screen "BC Max Step Times" 1280x800, template "Template"
   on GenerateScreen: "TitleUpdater"()
   Button "HmiScreenItemData_1" at 1,1 size 150x43; TextOn 'Back'; TextOff 'Commissioning'
      on Release: ActivateScreen("Commissioning Main Page", 0)
   Button "Button_1" at 21,736 size 161x32; TextOff 'Back'
      on Activate: ActivateScreen("IGG Process Times", 0)
   TextField "Text field_25" at 83,285 size 286x22; Text 'Step 040'
   TextField "Text field_29" at 383,118 size 77x20; Text 'Time (ms)'
   TextField "Text field_33" at 83,312 size 286x22; Text 'Step 050'
   IOField "I/O field_58" at 382,312 size 60x22; Authorization "Parameter Change"; FormatPattern s9999999999
      ProcessValue <- "86_Times_STEP_MAX_TIME_STP_050(1)"
   TextField "Text field_35" at 83,367 size 286x22; Text 'Step 070'
   TextField "Text field_65" at 83,144 size 286x22; Text 'Step 001'
   TextField "Text field_67" at 83,173 size 286x22; Text 'Step 005'
   TextField "Text field_69" at 83,200 size 286x22; Text 'Step 010'
   TextField "Text field_71" at 83,229 size 286x22; Text 'Step 020'
   TextField "Text field_73" at 83,257 size 286x22; Text 'Step 030'
   TextField "Text field_42" at 83,118 size 89x20; Text 'Description'
   IOField "I/O field_128" at 382,144 size 60x22; Authorization "Parameter Change"; FormatPattern s9999999999
      ProcessValue <- "86_Times_STEP_MAX_TIME_STP_001(1)"
   IOField "I/O field_133" at 382,173 size 60x22; Authorization "Parameter Change"; FormatPattern s9999999999
      ProcessValue <- "86_Times_STEP_MAX_TIME_STP_005(1)"
   IOField "I/O field_138" at 382,200 size 60x22; Authorization "Parameter Change"; FormatPattern s9999999999
      ProcessValue <- "86_Times_STEP_MAX_TIME_STP_010(1)"
   IOField "I/O field_148" at 382,257 size 60x22; Authorization "Parameter Change"; FormatPattern s9999999999
      ProcessValue <- "86_Times_STEP_MAX_TIME_STP_030(1)"
   IOField "I/O field_64" at 382,367 size 60x22; Authorization "Parameter Change"; FormatPattern s9999999999
      ProcessValue <- "86_Times_STEP_MAX_TIME_STP_070(1)"
   TextField "Text field_53" at 82,92 size 247x26; Text 'BC Maximum Step Times'
   IOField "I/O field_5" at 382,229 size 60x22; Authorization "Parameter Change"; FormatPattern s9999999999
      ProcessValue <- "86_Times_STEP_MAX_TIME_STP_020(1)"
   TextField "Text field_1" at 83,340 size 286x22; Text 'Step 060'
   IOField "I/O field_2" at 382,340 size 60x22; Authorization "Parameter Change"; FormatPattern s9999999999
      ProcessValue <- "86_Times_STEP_MAX_TIME_STP_060(1)"
   TextField "Text field_2" at 461,286 size 286x22; Text 'Step 240'
   TextField "Text field_3" at 750,119 size 77x20; Text 'Time (ms)'
   TextField "Text field_4" at 461,313 size 286x22; Text 'Step 250'
   IOField "I/O field_1" at 758,312 size 60x22; Authorization "Parameter Change"; FormatPattern s9999999999
      ProcessValue <- "86_Times_STEP_MAX_TIME_STP_250(1)"
   TextField "Text field_5" at 461,368 size 286x22; Text 'Step 270'
   TextField "Text field_6" at 461,145 size 286x22; Text 'Step 190'
   TextField "Text field_7" at 461,174 size 286x22; Text 'Step 200'
   TextField "Text field_8" at 461,201 size 286x22; Text 'Step 210'
   TextField "Text field_9" at 461,230 size 286x22; Text 'Step 220'
   TextField "Text field_10" at 461,258 size 286x22; Text 'Step 230'
   TextField "Text field_11" at 461,119 size 89x20; Text 'Description'
   IOField "I/O field_3" at 758,145 size 60x22; Authorization "Parameter Change"; FormatPattern s9999999999
      ProcessValue <- "86_Times_STEP_MAX_TIME_STP_190(1)"
   IOField "I/O field_4" at 758,174 size 60x22; Authorization "Parameter Change"; FormatPattern s9999999999
      ProcessValue <- "86_Times_STEP_MAX_TIME_STP_200(1)"
   IOField "I/O field_6" at 758,201 size 60x22; Authorization "Parameter Change"; FormatPattern s9999999999
      ProcessValue <- "86_Times_STEP_MAX_TIME_STP_210(1)"
   IOField "I/O field_8" at 758,258 size 60x22; Authorization "Parameter Change"; FormatPattern s9999999999
      ProcessValue <- "86_Times_STEP_MAX_TIME_STP_230(1)"
   IOField "I/O field_9" at 758,367 size 60x22; Authorization "Parameter Change"; FormatPattern s9999999999
      ProcessValue <- "86_Times_STEP_MAX_TIME_STP_270(1)"
   IOField "I/O field_10" at 758,230 size 60x22; Authorization "Parameter Change"; FormatPattern s9999999999
      ProcessValue <- "86_Times_STEP_MAX_TIME_STP_220(1)"
   TextField "Text field_13" at 461,341 size 286x22; Text 'Step 260'
   IOField "I/O field_11" at 758,340 size 60x22; Authorization "Parameter Change"; FormatPattern s9999999999
      ProcessValue <- "86_Times_STEP_MAX_TIME_STP_260(1)"
   TextField "Text field_14" at 83,398 size 286x22; Text 'Step 080'
   IOField "I/O field_12" at 382,398 size 60x22; Authorization "Parameter Change"; FormatPattern s9999999999
      ProcessValue <- "86_Times_STEP_MAX_TIME_STP_080(1)"
   TextField "Text field_15" at 83,426 size 286x22; Text 'Step 090'
   IOField "I/O field_13" at 382,426 size 60x22; Authorization "Parameter Change"; FormatPattern s9999999999
      ProcessValue <- "86_Times_STEP_MAX_TIME_STP_090(1)"
   TextField "Text field_16" at 83,453 size 286x22; Text 'Step 100'
   IOField "I/O field_14" at 382,453 size 60x22; Authorization "Parameter Change"; FormatPattern s9999999999
      ProcessValue <- "86_Times_STEP_MAX_TIME_STP_100(1)"
   IOField "I/O field_15" at 382,285 size 60x22; Authorization "Parameter Change"; FormatPattern s9999999999
      ProcessValue <- "86_Times_STEP_MAX_TIME_STP_040(1)"
   TextField "Text field_17" at 461,395 size 286x22; Text 'Step 280'
   IOField "I/O field_16" at 758,394 size 60x22; Authorization "Parameter Change"; FormatPattern s9999999999
      ProcessValue <- "86_Times_STEP_MAX_TIME_STP_280(1)"
   TextField "Text field_18" at 461,426 size 286x22; Text 'Step 290'
   IOField "I/O field_17" at 758,425 size 60x22; Authorization "Parameter Change"; FormatPattern s9999999999
      ProcessValue <- "86_Times_STEP_MAX_TIME_STP_290(1)"
   TextField "Text field_19" at 461,453 size 286x22; Text 'Step 300'
   IOField "I/O field_18" at 758,452 size 60x22; Authorization "Parameter Change"; FormatPattern s9999999999
      ProcessValue <- "86_Times_STEP_MAX_TIME_STP_300(1)"
   TextField "Text field_20" at 461,483 size 286x22; Text 'Step 310'
   IOField "I/O field_19" at 758,482 size 60x22; Authorization "Parameter Change"; FormatPattern s9999999999
      ProcessValue <- "86_Times_STEP_MAX_TIME_STP_310(1)"
   TextField "Text field_21" at 461,510 size 286x22; Text 'Step 320'
   IOField "I/O field_20" at 758,509 size 60x22; Authorization "Parameter Change"; FormatPattern s9999999999
      ProcessValue <- "86_Times_STEP_MAX_TIME_STP_320(1)"
   TextField "Text field_22" at 835,145 size 286x22; Text 'Step 390'
   IOField "I/O field_21" at 1130,144 size 60x22; Authorization "Parameter Change"; FormatPattern s9999999999
      ProcessValue <- "86_Times_STEP_MAX_TIME_STP_390(1)"
   TextField "Text field_23" at 835,118 size 89x20; Text 'Description'
   TextField "Text field_24" at 1122,119 size 77x20; Text 'Time (ms)'
   TextField "Text field_26" at 835,173 size 286x22; Text 'Step 400'
   IOField "I/O field_22" at 1130,172 size 60x22; Authorization "Parameter Change"; FormatPattern s9999999999
      ProcessValue <- "86_Times_STEP_MAX_TIME_STP_400(1)"
   TextField "Text field_27" at 835,200 size 286x22; Text 'Step 410'
   IOField "I/O field_23" at 1130,199 size 60x22; Authorization "Parameter Change"; FormatPattern s9999999999
      ProcessValue <- "86_Times_STEP_MAX_TIME_STP_410(1)"
   TextField "Text field_28" at 835,230 size 286x22; Text 'Step 420'
   IOField "I/O field_24" at 1130,229 size 60x22; Authorization "Parameter Change"; FormatPattern s9999999999
      ProcessValue <- "86_Times_STEP_MAX_TIME_STP_420(1)"
   TextField "Text field_30" at 835,257 size 286x22; Text 'Step 430'
   IOField "I/O field_25" at 1130,256 size 60x22; Authorization "Parameter Change"; FormatPattern s9999999999
      ProcessValue <- "86_Times_STEP_MAX_TIME_STP_430(1)"
   TextField "Text field_31" at 835,285 size 286x22; Text 'Step 440'
   IOField "I/O field_26" at 1130,284 size 60x22; Authorization "Parameter Change"; FormatPattern s9999999999
      ProcessValue <- "86_Times_STEP_MAX_TIME_STP_440(1)"
   TextField "Text field_32" at 835,312 size 286x22; Text 'Step 450'
   IOField "I/O field_27" at 1130,311 size 60x22; Authorization "Parameter Change"; FormatPattern s9999999999
      ProcessValue <- "86_Times_STEP_MAX_TIME_STP_450(1)"
   TextField "Text field_34" at 835,341 size 286x22; Text 'Step 460'
   IOField "I/O field_28" at 1130,340 size 60x22; Authorization "Parameter Change"; FormatPattern s9999999999
      ProcessValue <- "86_Times_STEP_MAX_TIME_STP_460(1)"
   TextField "Text field_36" at 835,369 size 286x22; Text 'Step 470'
   IOField "I/O field_29" at 1130,368 size 60x22; Authorization "Parameter Change"; FormatPattern s9999999999
      ProcessValue <- "86_Times_STEP_MAX_TIME_STP_470(1)"
   TextField "Text field_37" at 835,395 size 286x22; Text 'Step 480'
   IOField "I/O field_30" at 1130,394 size 60x22; Authorization "Parameter Change"; FormatPattern s9999999999
      ProcessValue <- "86_Times_STEP_MAX_TIME_STP_480(1)"
   TextField "Text field_38" at 835,426 size 286x22; Text 'Step 490'
   IOField "I/O field_31" at 1130,425 size 60x22; Authorization "Parameter Change"; FormatPattern s9999999999
      ProcessValue <- "86_Times_STEP_MAX_TIME_STP_490(1)"
   TextField "Text field_39" at 835,452 size 286x22; Text 'Step 500'
   IOField "I/O field_32" at 1130,451 size 60x22; Authorization "Parameter Change"; FormatPattern s9999999999
      ProcessValue <- "86_Times_STEP_MAX_TIME_STP_500(1)"
   TextField "Text field_40" at 835,482 size 286x22; Text 'Step 510'
   IOField "I/O field_33" at 1130,481 size 60x22; Authorization "Parameter Change"; FormatPattern s9999999999
      ProcessValue <- "86_Times_STEP_MAX_TIME_STP_510(1)"
   TextField "Text field_41" at 835,510 size 286x22; Text 'Step 520'
   IOField "I/O field_34" at 1130,509 size 60x22; Authorization "Parameter Change"; FormatPattern s9999999999
      ProcessValue <- "86_Times_STEP_MAX_TIME_STP_520(1)"
   IOField "I/O field_7" at 758,285 size 60x22; Authorization "Parameter Change"; FormatPattern s9999999999
      ProcessValue <- "86_Times_STEP_MAX_TIME_STP_240(1)"
   TextField "Text field_43" at 83,483 size 286x22; Text 'Step 110'
   IOField "I/O field_35" at 382,483 size 60x22; Authorization "Parameter Change"; FormatPattern s9999999999
      ProcessValue <- "86_Times_STEP_MAX_TIME_STP_110(1)"
   TextField "Text field_44" at 83,510 size 286x22; Text 'Step 120'
   IOField "I/O field_36" at 382,510 size 60x22; Authorization "Parameter Change"; FormatPattern s9999999999
      ProcessValue <- "86_Times_STEP_MAX_TIME_STP_120(1)"
   TextField "Text field_45" at 461,538 size 286x22; Text 'Step 330'
   IOField "I/O field_37" at 758,537 size 60x22; Authorization "Parameter Change"; FormatPattern s9999999999
      ProcessValue <- "86_Times_STEP_MAX_TIME_STP_330(1)"
   TextField "Text field_46" at 835,538 size 286x22; Text 'Step 530'
   IOField "I/O field_38" at 1130,537 size 60x22; Authorization "Parameter Change"; FormatPattern s9999999999
      ProcessValue <- "86_Times_STEP_MAX_TIME_STP_530(1)"
   TextField "Text field_47" at 83,538 size 286x22; Text 'Step 130'
   IOField "I/O field_39" at 382,538 size 60x22; Authorization "Parameter Change"; FormatPattern s9999999999
      ProcessValue <- "86_Times_STEP_MAX_TIME_STP_130(1)"
   TextField "Text field_48" at 461,568 size 286x22; Text 'Step 340'
   IOField "I/O field_40" at 758,567 size 60x22; Authorization "Parameter Change"; FormatPattern s9999999999
      ProcessValue <- "86_Times_STEP_MAX_TIME_STP_340(1)"
   TextField "Text field_49" at 835,568 size 286x22; Text 'Step 540'
   IOField "I/O field_41" at 1130,567 size 60x22; Authorization "Parameter Change"; FormatPattern s9999999999
      ProcessValue <- "86_Times_STEP_MAX_TIME_STP_540(1)"
   TextField "Text field_50" at 83,568 size 286x22; Text 'Step 140'
   IOField "I/O field_42" at 382,568 size 60x22; Authorization "Parameter Change"; FormatPattern s9999999999
      ProcessValue <- "86_Times_STEP_MAX_TIME_STP_140(1)"
   TextField "Text field_51" at 461,599 size 286x22; Text 'Step 350'
   IOField "I/O field_43" at 758,598 size 60x22; Authorization "Parameter Change"; FormatPattern s9999999999
      ProcessValue <- "86_Times_STEP_MAX_TIME_STP_350(1)"
   TextField "Text field_52" at 835,599 size 286x22; Text 'Step 550'
   IOField "I/O field_44" at 1130,598 size 60x22; Authorization "Parameter Change"; FormatPattern s9999999999
      ProcessValue <- "86_Times_STEP_MAX_TIME_STP_550(1)"
   TextField "Text field_54" at 83,599 size 286x22; Text 'Step 150'
   IOField "I/O field_45" at 382,599 size 60x22; Authorization "Parameter Change"; FormatPattern s9999999999
      ProcessValue <- "86_Times_STEP_MAX_TIME_STP_150(1)"
   TextField "Text field_55" at 461,628 size 286x22; Text 'Step 360'
   IOField "I/O field_46" at 758,627 size 60x22; Authorization "Parameter Change"; FormatPattern s9999999999
      ProcessValue <- "86_Times_STEP_MAX_TIME_STP_360(1)"
   TextField "Text field_56" at 835,628 size 286x22; Text 'Step 560'
   IOField "I/O field_47" at 1130,627 size 60x22; Authorization "Parameter Change"; FormatPattern s9999999999
      ProcessValue <- "86_Times_STEP_MAX_TIME_STP_560(1)"
   TextField "Text field_57" at 83,628 size 286x22; Text 'Step 160'
   IOField "I/O field_48" at 382,628 size 60x22; Authorization "Parameter Change"; FormatPattern s9999999999
      ProcessValue <- "86_Times_STEP_MAX_TIME_STP_160(1)"
   TextField "Text field_58" at 461,657 size 286x22; Text 'Step 370'
   IOField "I/O field_49" at 758,656 size 60x22; Authorization "Parameter Change"; FormatPattern s9999999999
      ProcessValue <- "86_Times_STEP_MAX_TIME_STP_370(1)"
   TextField "Text field_59" at 835,657 size 286x22; Text 'Step 570'
   IOField "I/O field_50" at 1130,656 size 60x22; Authorization "Parameter Change"; FormatPattern s9999999999
      ProcessValue <- "86_Times_STEP_MAX_TIME_STP_570(1)"
   TextField "Text field_60" at 83,657 size 286x22; Text 'Step 170'
   IOField "I/O field_51" at 382,657 size 60x22; Authorization "Parameter Change"; FormatPattern s9999999999
      ProcessValue <- "86_Times_STEP_MAX_TIME_STP_170(1)"
   TextField "Text field_61" at 461,687 size 286x22; Text 'Step 380'
   IOField "I/O field_52" at 758,686 size 60x22; Authorization "Parameter Change"; FormatPattern s9999999999
      ProcessValue <- "86_Times_STEP_MAX_TIME_STP_380(1)"
   TextField "Text field_63" at 83,687 size 286x22; Text 'Step 180'
   IOField "I/O field_54" at 382,687 size 60x22; Authorization "Parameter Change"; FormatPattern s9999999999
      ProcessValue <- "86_Times_STEP_MAX_TIME_STP_180(1)"
   Group "Group" at 455,41 size 373x50
   Button "HmiScreenItemData_8" at 469,45 size 355x40; TextOn 'Back'; TextOff 'Text'
   TextField "Screen title" at 455,41 size 373x50; Text 'Screen title'

screen "BC Digital Inputs" 1280x800, template "Template"
   on GenerateScreen: "TitleUpdater"()
   Button "HmiScreenItemData_1" at 1,1 size 150x43; TextOn 'Back'; TextOff 'Commissioning'
      on Release: ActivateScreen("Commissioning Main Page", 0)
   TextField "Text field_37" at 361,69 size 287x26; Text 'Burner Control PLC (Rack 2)'
   TextField "Text field_38" at 361,139 size 55x22; Text 'I0.0'
   TextField "Text field_39" at 361,174 size 55x22; Text 'I0.1'
   TextField "Text field_40" at 361,210 size 55x22; Text 'I0.2'
   TextField "Text field_41" at 361,246 size 55x22; Text 'I0.3'
   TextField "Text field_42" at 361,282 size 55x22; Text 'I0.4'
   TextField "Text field_43" at 361,318 size 55x22; Text 'I0.5'
   TextField "Text field_44" at 361,354 size 55x22; Text 'I0.6'
   TextField "Text field_45" at 361,390 size 55x22; Text 'I0.7'
   Circle "Circle_33" at 421,139 size 20x20
      Appearance <- "10 DI_DATA_PS101"
   Circle "Circle_34" at 421,175 size 20x20
      Appearance <- "10 DI_DATA_E131_SHTDN"
   Circle "Circle_35" at 421,211 size 20x20
      Appearance <- "10 DI_DATA_R2_SPR_DI_0_2"
   Circle "Circle_36" at 421,247 size 20x20
      Appearance <- "10 DI_DATA_R2_SPR_DI_0_3"
   Circle "Circle_37" at 421,282 size 20x20
      Appearance <- "10 DI_DATA_X001_PWR_OK"
   Circle "Circle_38" at 421,318 size 20x20
      Appearance <- "10 DI_DATA_FD001_PWR_OK"
   Circle "Circle_39" at 421,354 size 20x20
      Appearance <- "10 DI_DATA_FD001_OK"
   Circle "Circle_40" at 421,390 size 20x20
      Appearance <- "103_Main_Burner_DB_DN_OK(1)"
   TextField "Text field_46" at 378,107 size 49x26; Text 'I0'
   TextField "Text field_47" at 361,458 size 55x22; Text 'I1.0'
   TextField "Text field_48" at 361,493 size 55x22; Text 'I1.1'
   TextField "Text field_49" at 361,529 size 55x22; Text 'I1.2'
   TextField "Text field_50" at 361,565 size 55x22; Text 'I1.3'
   TextField "Text field_51" at 361,601 size 55x22; Text 'I1.4'
   TextField "Text field_52" at 361,637 size 55x22; Text 'I1.5'
   TextField "Text field_53" at 361,673 size 55x22; Text 'I1.6'
   TextField "Text field_54" at 361,709 size 55x22; Text 'I1.7'
   Circle "Circle_41" at 421,458 size 20x20
      Appearance <- "10 DI_DATA_FS123"
   Circle "Circle_42" at 421,494 size 20x20
      Appearance <- "10 DI_DATA_FS115(1)"
   Circle "Circle_43" at 421,530 size 20x20
      Appearance <- "10 DI_DATA_FS320"
   Circle "Circle_44" at 421,566 size 20x20
      Appearance <- "10 DI_DATA_FS317"
   Circle "Circle_45" at 421,601 size 20x20
      Appearance <- "10 DI_DATA_P301_TRIPPED(1)"
   Circle "Circle_46" at 421,637 size 20x20
      Appearance <- "10 DI_DATA_P301_ENBLD"
   Circle "Circle_47" at 421,673 size 20x20
      Appearance <- "10 DI_DATA_R2_SPR_DI_1_6"
   Circle "Circle_48" at 421,709 size 20x20
      Appearance <- "10 DI_DATA_ESD_OK"
   TextField "Text field_55" at 378,426 size 49x26; Text 'I1'
   TextField "Text field_56" at 652,139 size 55x22; Text 'I2.0'
   TextField "Text field_57" at 652,174 size 55x22; Text 'I2.1'
   TextField "Text field_58" at 652,210 size 55x22; Text 'I2.2'
   TextField "Text field_59" at 652,246 size 55x22; Text 'I2.3'
   TextField "Text field_60" at 652,282 size 55x22; Text 'I2.4'
   TextField "Text field_61" at 652,318 size 55x22; Text 'I2.5'
   TextField "Text field_62" at 652,354 size 55x22; Text 'I2.6'
   TextField "Text field_63" at 652,390 size 55x22; Text 'I2.7'
   Circle "Circle_49" at 712,139 size 20x20
      Appearance <- "10 DI_DATA_E600_NOK"
   Circle "Circle_50" at 712,175 size 20x20
      Appearance <- "10 DI_DATA_E600_HIHI"
   Circle "Circle_51" at 712,211 size 20x20
      Appearance <- "10 DI_DATA_E600_LOLO"
   Circle "Circle_52" at 712,247 size 20x20
      Appearance <- "10 DI_DATA_E600_PWR_OK"
   Circle "Circle_53" at 712,282 size 20x20
      Appearance <- "10 DI_DATA_E700_PWR_OK"
   Circle "Circle_54" at 712,318 size 20x20
      Appearance <- "10 DI_DATA_E700_OPACITY"
   Circle "Circle_55" at 712,354 size 20x20
      Appearance <- "10 DI_DATA_TS403_FAULT(1)"
   Circle "Circle_56" at 712,390 size 20x20
      Appearance <- "10 DI_DATA_TS006"
   TextField "Text field_64" at 669,107 size 49x26; Text 'I2'
   TextField "Text field_65" at 650,458 size 55x22; Text 'I3.0'
   TextField "Text field_66" at 650,493 size 55x22; Text 'I3.1'
   TextField "Text field_67" at 650,529 size 55x22; Text 'I3.2'
   TextField "Text field_68" at 650,565 size 55x22; Text 'I3.3'
   TextField "Text field_69" at 650,601 size 55x22; Text 'I3.4'
   TextField "Text field_70" at 650,637 size 55x22; Text 'I3.5'
   TextField "Text field_71" at 650,673 size 55x22; Text 'I3.6'
   TextField "Text field_72" at 650,709 size 55x22; Text 'I3.7'
   Circle "Circle_57" at 710,458 size 20x20
      Appearance <- "10 DI_DATA_S2_8K1_OK"
   Circle "Circle_58" at 710,494 size 20x20
      Appearance <- "10 DI_DATA_E131_WRNG"
   Circle "Circle_59" at 710,530 size 20x20
      Appearance <- "10 DI_DATA_R2_SPR_DI_3_2"
   Circle "Circle_60" at 710,566 size 20x20
      Appearance <- "10 DI_DATA_E131_OK"
   Circle "Circle_61" at 710,601 size 20x20
      Appearance <- "10 DI_DATA_LS001"
   Circle "Circle_62" at 710,637 size 20x20
      Appearance <- "10 DI_DATA_P305_TRIPPED"
   Circle "Circle_63" at 710,673 size 20x20
      Appearance <- "10 DI_DATA_P305_ENBLD"
   Circle "Circle_64" at 710,709 size 20x20
      Appearance <- "10 DI_DATA_R2_SPR_DI_3_7"
   TextField "Text field_73" at 667,426 size 49x26; Text 'I3'
   TextField "Text field_107" at 450,138 size 180x22; Text 'CA Pressure Switch PS101'
   TextField "Text field_108" at 450,176 size 180x22; Text 'IA Comp Shutdown E131'
   TextField "Text field_109" at 449,216 size 180x22; Text 'Spare Input'
   TextField "Text field_110" at 449,250 size 180x22; Text 'Spare Input'
   TextField "Text field_111" at 449,282 size 180x22; Text 'Ignitor Power Healthy X001'
   TextField "Text field_112" at 449,317 size 180x22; Text 'FDU Power Healthy FD001'
   TextField "Text field_113" at 449,353 size 180x22; Text 'FDU Healthy FD001'
   TextField "Text field_114" at 449,390 size 180x22; Text 'Burner Flame Detected FD001'
   TextField "Text field_116" at 447,458 size 180x22; Text 'Pilot Ign. Air Flow Sw FS123'
   TextField "Text field_117" at 447,494 size 180x22; Text 'Main Atom Air Flow Sw FS115'
   TextField "Text field_118" at 447,529 size 180x22; Text 'Nozzle CW Flow Sw FS320'
   TextField "Text field_119" at 447,566 size 180x22; Text 'Jacket CW Flow Sw FS317'
   TextField "Text field_120" at 447,602 size 180x22; Text 'CSW Pump Tripped P301'
   TextField "Text field_121" at 447,637 size 180x22; Text 'CSW Pump Enabled P301'
   TextField "Text field_122" at 447,710 size 180x22; Text 'Ext. Shutdown'
   TextField "Text field_123" at 740,137 size 180x22; Text 'O2 System Fail E600'
   TextField "Text field_124" at 740,174 size 180x22; Text 'O2 Hi Hi E600'
   TextField "Text field_125" at 739,210 size 180x22; Text 'O2 Lo Lo E600'
   TextField "Text field_126" at 739,246 size 180x22; Text 'O2 System Power Healthy E600'
   TextField "Text field_127" at 739,280 size 180x22; Text 'Soot System Power Healthy E700'
   TextField "Text field_128" at 739,315 size 180x22; Text 'Soot System Opacity E700'
   TextField "Text field_129" at 739,352 size 180x22; Text 'IG Temp Hi Hi Switch TS403'
   TextField "Text field_130" at 740,390 size 180x22; Text 'IG Shell Temp Hi Switch TS006'
   TextField "Text field_131" at 739,458 size 180x22; Text 'IGG E-Stop Healthy'
   TextField "Text field_132" at 739,493 size 180x22; Text 'IA Comp Warning E131'
   TextField "Text field_133" at 739,529 size 180x22; Text 'Spare Input'
   TextField "Text field_134" at 739,637 size 180x22; Text 'Fresh Water Pump Tripped P305'
   TextField "Text field_135" at 739,673 size 180x22; Text 'Fresh Water Pump Enabled P305'
   TextField "Text field_136" at 739,709 size 180x22; Text 'Spare Input'
   TextField "Text field_137" at 739,565 size 180x22; Text 'IA Comp Healthy E131'
   TextField "Text field_138" at 739,601 size 180x22; Text 'Shell CW Level Hi Hi Sw LS001'
   TextField "Text field_115" at 447,673 size 180x22; Text 'Spare Input'
   Group "Group" at 740,44 size 373x50
   Button "HmiScreenItemData_8" at 754,48 size 355x40; TextOn 'Back'; TextOff 'Text'
   TextField "Screen title" at 740,44 size 373x50; Text 'Screen title'

screen "GCU Digital Inputs" 1280x800, template "Template"
   on GenerateScreen: "TitleUpdater"()
   Button "HmiScreenItemData_1" at 1,1 size 150x43; TextOn 'Back'; TextOff 'Commissioning'
      on Release: ActivateScreen("Commissioning Main Page", 0)
   AlarmView "Alarm view_1" at 0,777 size 1280x23
   TextField "Text field_37" at 165,44 size 300x30; Text 'GCU Control PLC (Rack 3)'
   TextField "Text field_34" at 745,74 size 60x30; Text 'I 2'
   TextField "Text field_35" at 745,384 size 70x22; Text 'I 138.7'
   Circle "Circle_16" at 825,384 size 20x20
      Appearance <- "10_DI_DATA_P_303_ENBLD"
   TextField "Text field_36" at 865,384 size 230x22; Text 'P303 ENABLED'
   TextField "Text field_39" at 745,344 size 70x22; Text 'I 138.6'
   Circle "Circle_17" at 825,344 size 20x20
      Appearance <- "10_DI_DATA_EPB_8S1"
   TextField "Text field_40" at 865,344 size 230x22; Text 'PB E-STOP'
   TextField "Text field_41" at 745,304 size 70x22; Text 'I 138.5'
   Circle "Circle_18" at 825,304 size 20x20
      Appearance <- "10_DI_DATA_PB_10S2"
   TextField "Text field_42" at 865,304 size 230x22; Text 'PB STOP'
   TextField "Text field_43" at 745,264 size 70x22; Text 'I 138.4'
   Circle "Circle_19" at 825,264 size 20x20
      Appearance <- "10_DI_DATA_PB_10S1"
   TextField "Text field_44" at 865,264 size 230x22; Text 'PB START'
   TextField "Text field_45" at 745,224 size 70x22; Text 'I 138.3'
   Circle "Circle_20" at 825,224 size 20x20
      Appearance <- "10_DI_DATA_P_304_ENBLD"
   TextField "Text field_46" at 865,224 size 230x22; Text 'P304 ENABLED'
   TextField "Text field_47" at 745,184 size 70x22; Text 'I 138.2'
   Circle "Circle_21" at 825,184 size 20x20
      Appearance <- "10_DI_DATA_LS_303_LO"
   TextField "Text field_48" at 863,184 size 230x22; Text 'LS303 GCU LOW LEVEL'
   TextField "Text field_49" at 745,144 size 70x22; Text 'I 138.1'
   Circle "Circle_22" at 825,144 size 20x20
      Appearance <- "10_DI_DATA_CV441_CLSD"
   TextField "Text field_50" at 865,144 size 230x22; Text 'CV441 CLOSED'
   TextField "Text field_51" at 745,104 size 70x22; Text 'I 138.0'
   Circle "Circle_23" at 825,104 size 20x20
      Appearance <- "10_DI_DATA_CV441_OPN"
   TextField "Text field_52" at 865,104 size 230x22; Text 'CV441 OPEN'
   TextField "Text field_53" at 745,424 size 60x30; Text 'I 3'
   TextField "Text field_54" at 745,734 size 70x22; Text 'I 139.7'
   Circle "Circle_24" at 825,734 size 20x20
      Appearance <- "10_DI_DATA_E_400_NOK"
   TextField "Text field_55" at 865,734 size 230x22; Text 'E400 FAULT'
   TextField "Text field_56" at 745,694 size 70x22; Text 'I 139.6'
   Circle "Circle_25" at 825,694 size 20x20
      Appearance <- "10_DI_DATA_E_400_RUN"
   TextField "Text field_57" at 865,694 size 230x22; Text 'E400 LOADED'
   TextField "Text field_58" at 745,654 size 70x22; Text 'I 139.5'
   Circle "Circle_26" at 825,654 size 20x20
      Appearance <- "10_DI_DATA_P_304_OK"
   TextField "Text field_59" at 865,654 size 230x22; Text 'P304 HEALTHY'
   TextField "Text field_60" at 745,614 size 70x22; Text 'I 139.4'
   Circle "Circle_27" at 825,614 size 20x20
      Appearance <- "10_DI_DATA_6Q6_PWR_OK"
   TextField "Text field_61" at 865,614 size 230x22; Text 'PANEL VENT POWER OK'
   TextField "Text field_62" at 745,574 size 70x22; Text 'I 139.3'
   Circle "Circle_28" at 825,574 size 20x20
      Appearance <- "10_DI_DATA_5T1_PWR_OK"
   TextField "Text field_63" at 865,574 size 230x22; Text '5T1 POWER OK'
   TextField "Text field_64" at 745,534 size 70x22; Text 'I 139.2'
   Circle "Circle_29" at 825,534 size 20x20
      Appearance <- "10_DI_DATA_P_303_OK"
   TextField "Text field_65" at 865,534 size 230x22; Text 'P303 HEALTHY'
   TextField "Text field_66" at 745,494 size 70x22; Text 'I 139.1'
   Circle "Circle_30" at 825,494 size 20x20
      Appearance <- "10_DI_DATA_E_400_SHTDN"
   TextField "Text field_67" at 865,494 size 230x22; Text 'E400 TRIPPED / FAULT'
   TextField "Text field_68" at 745,454 size 70x22; Text 'I 139.0'
   Circle "Circle_31" at 825,454 size 20x20
      Appearance <- "Process Gas Compressor Running/Stopped"
   TextField "Text field_69" at 865,454 size 230x22; Text 'E400 RUN / STOP'
   TextField "Text field_1" at 165,74 size 60x30; Text 'I 0'
   TextField "Text field_15" at 165,384 size 70x22; Text 'I 136.7'
   Circle "Circle_7" at 245,384 size 20x20
      Appearance <- "10_DI_DATA_CV341_CLSD"
   TextField "Text field_16" at 285,384 size 230x22; Text 'CV341 CLOSED'
   TextField "Text field_13" at 165,344 size 70x22; Text 'I 136.6'
   Circle "Circle_6" at 245,344 size 20x20
      Appearance <- "10_DI_DATA_CV341_OPN"
   TextField "Text field_14" at 285,344 size 230x22; Text 'CV341 OPEN'
   TextField "Text field_11" at 165,304 size 70x22; Text 'I 136.5'
   Circle "Circle_5" at 245,304 size 20x20
      Appearance <- "10_DI_DATA_FS_350_FLW_OK"
   TextField "Text field_12" at 285,304 size 230x22; Text 'FS350 FCW FLOW'
   TextField "Text field_9" at 165,264 size 70x22; Text 'I 136.4'
   Circle "Circle_4" at 245,264 size 20x20
      Appearance <- "10_DI_DATA_CV358_CLSD"
   TextField "Text field_10" at 285,264 size 230x22; Text 'CV358 CLOSED'
   TextField "Text field_7" at 165,224 size 70x22; Text 'I 136.3'
   Circle "Circle_3" at 245,224 size 20x20
      Appearance <- "10_DI_DATA_CV358_OPN"
   TextField "Text field_8" at 285,224 size 230x22; Text 'CV358 OPEN'
   TextField "Text field_5" at 165,184 size 70x22; Text 'I 136.2'
   Circle "Circle_2" at 245,184 size 20x20
      Appearance <- "10_DI_DATA_FS_332 FLW_OK"
   TextField "Text field_6" at 285,184 size 230x22; Text 'FS332 CSW FLOW'
   TextField "Text field_3" at 165,144 size 70x22; Text 'I 136.1'
   Circle "Circle_1" at 245,144 size 20x20
      Appearance <- "10_DI_DATA_R3_SPR_DI_136_1"
   TextField "Text field_4" at 285,144 size 230x22; Text 'R3_SPR_DI_136_1'
   TextField "Text field_38" at 165,104 size 70x22; Text 'I 136.0'
   Circle "Circle_33" at 245,104 size 20x20
      Appearance <- "10_DI_DATA_R3_SPR_DI_136_0"
   TextField "Text field_2" at 285,104 size 230x22; Text 'R3_SPR_DI_136_0'
   TextField "Text field_17" at 165,424 size 60x30; Text 'I 1'
   TextField "Text field_18" at 165,734 size 70x22; Text 'I 137.7'
   Circle "Circle_8" at 245,734 size 20x20
      Appearance <- "10_DI_DATA_CV409_CLSD"
   TextField "Text field_19" at 285,734 size 230x22; Text 'CV409 CLOSED'
   TextField "Text field_20" at 165,694 size 70x22; Text 'I 137.6'
   Circle "Circle_9" at 245,694 size 20x20
      Appearance <- "10_DI_DATA_CV409_OPN"
   TextField "Text field_21" at 285,694 size 230x22; Text 'CV409 OPEN'
   TextField "Text field_22" at 165,654 size 70x22; Text 'I 137.5'
   Circle "Circle_10" at 245,654 size 20x20
      Appearance <- "10_DI_DATA_CV411_CLSD"
   TextField "Text field_23" at 285,654 size 230x22; Text 'CV411 CLOSED'
   TextField "Text field_24" at 165,614 size 70x22; Text 'I 137.4'
   Circle "Circle_11" at 245,614 size 20x20
      Appearance <- "10_DI_DATA_CV411_OPN"
   TextField "Text field_25" at 285,614 size 230x22; Text 'CV411 OPEN'
   TextField "Text field_26" at 165,574 size 70x22; Text 'I 137.3'
   Circle "Circle_12" at 245,574 size 20x20
      Appearance <- "10_DI_DATA_CV407_CLSD"
   TextField "Text field_27" at 285,574 size 230x22; Text 'CV407 CLOSED'
   TextField "Text field_28" at 165,534 size 70x22; Text 'I 137.2'
   Circle "Circle_13" at 245,534 size 20x20
      Appearance <- "10_DI_DATA_CV407_OPN"
   TextField "Text field_29" at 285,534 size 230x22; Text 'CV407 OPEN'
   TextField "Text field_30" at 165,494 size 70x22; Text 'I 137.1'
   Circle "Circle_14" at 245,494 size 20x20
      Appearance <- "10_DI_DATA_CV406_CLSD"
   TextField "Text field_31" at 285,494 size 230x22; Text 'CV406 CLOSED'
   TextField "Text field_32" at 165,454 size 70x22; Text 'I 137.0'
   Circle "Circle_15" at 245,454 size 20x20
      Appearance <- "10_DI_DATA_CV406_OPN"
   TextField "Text field_33" at 285,454 size 230x22; Text 'CV406 OPEN'
   Group "Group_1" at 851,41 size 373x50
   Button "HmiScreenItemData_8" at 865,45 size 355x40; TextOn 'Back'; TextOff 'Text'
   TextField "Screen title" at 851,41 size 373x50; Text 'Screen title'

screen "BWT Digital Inputs" 1280x800, template "Template"
   on GenerateScreen: "TitleUpdater"()
   TextField "Text field_37" at 16,52 size 263x26; Text 'BWT Control PLC (Rack 3)'
   TextField "Text field_38" at 16,122 size 55x22; Text 'I0.0'
   TextField "Text field_39" at 16,158 size 55x22; Text 'I0.1'
   TextField "Text field_40" at 16,194 size 55x22; Text 'I0.2'
   TextField "Text field_41" at 16,230 size 55x22; Text 'I0.3'
   TextField "Text field_42" at 16,265 size 55x22; Text 'I0.4'
   TextField "Text field_43" at 16,301 size 55x22; Text 'I0.5'
   TextField "Text field_44" at 16,337 size 55x22; Text 'I0.6'
   TextField "Text field_45" at 16,373 size 55x22; Text 'I0.7'
   Circle "Circle_33" at 76,122 size 20x20
      Appearance <- "10 DI_DATA_PS101"
   Circle "Circle_34" at 76,158 size 20x20
      Appearance <- "10 DI_DATA_E131_SHTDN"
   Circle "Circle_35" at 76,194 size 20x20
      Appearance <- "10 DI_DATA_R2_SPR_DI_0_2"
   Circle "Circle_36" at 76,230 size 20x20
      Appearance <- "10 DI_DATA_R2_SPR_DI_0_3"
   Circle "Circle_37" at 76,265 size 20x20
      Appearance <- "10 DI_DATA_X001_PWR_OK"
   Circle "Circle_38" at 76,301 size 20x20
      Appearance <- "10 DI_DATA_FD001_PWR_OK"
   Circle "Circle_39" at 76,337 size 20x20
      Appearance <- "10 DI_DATA_FD001_OK"
   Circle "Circle_40" at 76,373 size 20x20
      Appearance <- "103_Main_Burner_DB_DN_OK(1)"
   TextField "Text field_46" at 33,90 size 49x26; Text 'I0'
   TextField "Text field_47" at 16,441 size 55x22; Text 'I1.0'
   TextField "Text field_48" at 16,477 size 55x22; Text 'I1.1'
   TextField "Text field_49" at 16,513 size 55x22; Text 'I1.2'
   TextField "Text field_50" at 16,549 size 55x22; Text 'I1.3'
   TextField "Text field_51" at 16,584 size 55x22; Text 'I1.4'
   TextField "Text field_52" at 16,620 size 55x22; Text 'I1.5'
   TextField "Text field_53" at 16,656 size 55x22; Text 'I1.6'
   TextField "Text field_54" at 16,692 size 55x22; Text 'I1.7'
   Circle "Circle_41" at 76,441 size 20x20
      Appearance <- "10 DI_DATA_FS123"
   Circle "Circle_42" at 76,477 size 20x20
      Appearance <- "10 DI_DATA_FS115(1)"
   Circle "Circle_43" at 76,513 size 20x20
      Appearance <- "10 DI_DATA_FS320"
   Circle "Circle_44" at 76,549 size 20x20
      Appearance <- "10 DI_DATA_FS317"
   Circle "Circle_45" at 76,584 size 20x20
      Appearance <- "10 DI_DATA_P301_TRIPPED(1)"
   Circle "Circle_46" at 76,620 size 20x20
      Appearance <- "10 DI_DATA_P301_ENBLD"
   Circle "Circle_47" at 76,656 size 20x20
      Appearance <- "10 DI_DATA_R2_SPR_DI_1_6"
   Circle "Circle_48" at 76,692 size 20x20
      Appearance <- "10 DI_DATA_ESD_OK"
   TextField "Text field_55" at 33,409 size 49x26; Text 'I1'
   TextField "Text field_56" at 307,122 size 55x22; Text 'I2.0'
   TextField "Text field_57" at 307,158 size 55x22; Text 'I2.1'
   TextField "Text field_58" at 307,194 size 55x22; Text 'I2.2'
   TextField "Text field_59" at 307,230 size 55x22; Text 'I2.3'
   TextField "Text field_60" at 307,265 size 55x22; Text 'I2.4'
   TextField "Text field_61" at 307,301 size 55x22; Text 'I2.5'
   TextField "Text field_62" at 307,337 size 55x22; Text 'I2.6'
   TextField "Text field_63" at 307,373 size 55x22; Text 'I2.7'
   Circle "Circle_49" at 367,122 size 20x20
      Appearance <- "10 DI_DATA_E600_NOK"
   Circle "Circle_50" at 367,158 size 20x20
      Appearance <- "10 DI_DATA_E600_HIHI"
   Circle "Circle_51" at 367,194 size 20x20
      Appearance <- "10 DI_DATA_E600_LOLO"
   Circle "Circle_52" at 367,230 size 20x20
      Appearance <- "10 DI_DATA_E600_PWR_OK"
   Circle "Circle_53" at 367,265 size 20x20
      Appearance <- "10 DI_DATA_E700_PWR_OK"
   Circle "Circle_54" at 367,301 size 20x20
      Appearance <- "10 DI_DATA_E700_OPACITY"
   Circle "Circle_55" at 367,337 size 20x20
      Appearance <- "10 DI_DATA_TS403_FAULT(1)"
   Circle "Circle_56" at 367,373 size 20x20
      Appearance <- "10 DI_DATA_TS006"
   TextField "Text field_64" at 324,90 size 49x26; Text 'I2'
   TextField "Text field_65" at 305,441 size 46x22; Text 'I3.0'
   TextField "Text field_66" at 305,477 size 46x22; Text 'I3.1'
   TextField "Text field_67" at 305,513 size 46x22; Text 'I3.2'
   TextField "Text field_68" at 305,549 size 46x22; Text 'I3.3'
   TextField "Text field_69" at 305,584 size 46x22; Text 'I3.4'
   TextField "Text field_70" at 305,620 size 46x22; Text 'I3.5'
   TextField "Text field_71" at 305,656 size 46x22; Text 'I3.6'
   TextField "Text field_72" at 305,692 size 46x22; Text 'I3.7'
   Circle "Circle_57" at 365,441 size 20x20
      Appearance <- "10 DI_DATA_S2_8K1_OK"
   Circle "Circle_58" at 365,477 size 20x20
      Appearance <- "10 DI_DATA_E131_WRNG"
   Circle "Circle_59" at 365,513 size 20x20
      Appearance <- "10 DI_DATA_R2_SPR_DI_3_2"
   Circle "Circle_60" at 365,549 size 20x20
      Appearance <- "10 DI_DATA_E131_OK"
   Circle "Circle_61" at 365,584 size 20x20
      Appearance <- "10 DI_DATA_LS001"
   Circle "Circle_62" at 365,620 size 20x20
      Appearance <- "10 DI_DATA_P305_TRIPPED"
   Circle "Circle_63" at 365,656 size 20x20
      Appearance <- "10 DI_DATA_P305_ENBLD"
   Circle "Circle_64" at 365,692 size 20x20
      Appearance <- "10 DI_DATA_R2_SPR_DI_3_7"
   TextField "Text field_73" at 322,409 size 49x26; Text 'I3'
   Button "HmiScreenItemData_1" at 1,1 size 150x43; TextOn 'Back'; TextOff 'Commissioning'
      on Release: ActivateScreen("Commissioning Main Page", 0)
   TextField "Text field_107" at 105,111 size 243x23; Text 'CA Pressure Switch PS101'
   TextField "Text field_108" at 105,151 size 227x23; Text 'IA Comp Shutdown E131'
   TextField "Text field_109" at 104,191 size 112x23; Text 'Spare Input'
   TextField "Text field_110" at 104,225 size 112x23; Text 'Spare Input'
   TextField "Text field_111" at 104,257 size 258x23; Text 'Ignitor Power Healthy X001'
   TextField "Text field_112" at 104,292 size 181x42; Text 'FDU Power Healthy FD001'
   TextField "Text field_113" at 104,328 size 118x42; Text 'FDU Healthy FD001'
   TextField "Text field_114" at 104,365 size 215x42; Text 'Burner Flame Detected FD001'
   TextField "Text field_116" at 102,432 size 204x42; Text 'Pilot Ign. Air Flow Sw FS123'
   TextField "Text field_117" at 101,468 size 216x42; Text 'Main Atom Air Flow Sw FS115'
   TextField "Text field_118" at 101,504 size 182x42; Text 'Nozzle CW Flow Sw FS320'
   TextField "Text field_119" at 102,541 size 180x42; Text 'Jacket CW Flow Sw FS317'
   TextField "Text field_120" at 102,576 size 178x42; Text 'CSW Pump Tripped P301'
   TextField "Text field_121" at 105,611 size 180x42; Text 'CSW Pump Enabled P301'
   TextField "Text field_122" at 103,690 size 136x23; Text 'Ext. Shutdown'
   TextField "Text field_123" at 395,113 size 140x42; Text 'O2 System Fail E600'
   TextField "Text field_124" at 395,150 size 80x42; Text 'O2 Hi Hi E600'
   TextField "Text field_125" at 394,186 size 84x42; Text 'O2 Lo Lo E600'
   TextField "Text field_126" at 394,222 size 240x42; Text 'O2 System Power Healthy E600'
   TextField "Text field_127" at 394,256 size 257x42; Text 'Soot System Power Healthy E700'
   TextField "Text field_128" at 394,291 size 192x42; Text 'Soot System Opacity E700'
   TextField "Text field_129" at 394,328 size 199x42; Text 'IG Temp Hi Hi Switch TS403'
   TextField "Text field_130" at 395,366 size 225x42; Text 'IG Shell Temp Hi Switch TS006'
   TextField "Text field_131" at 394,437 size 181x23; Text 'IGG E-Stop Healthy'
   TextField "Text field_132" at 394,468 size 164x42; Text 'IA Comp Warning E131'
   TextField "Text field_133" at 393,509 size 112x23; Text 'Spare Input'
   TextField "Text field_134" at 393,611 size 248x42; Text 'Fresh Water Pump Tripped P305'
   TextField "Text field_135" at 393,648 size 250x42; Text 'Fresh Water Pump Enabled P305'
   TextField "Text field_136" at 394,688 size 112x23; Text 'Spare Input'
   TextField "Text field_137" at 395,540 size 159x42; Text 'IA Comp Healthy E131'
   TextField "Text field_138" at 394,576 size 222x42; Text 'Shell CW Level Hi Hi Sw LS001'
   TextField "Text field_115" at 105,654 size 112x23; Text 'Spare Input'
   AlarmView "Alarm view_1" at 0,777 size 1280x23
   TextField "Text field_1" at 23,309 size 1188x123; Text 'Re - Work Required Througout This page'
   Group "Group" at 455,41 size 373x50
   Button "HmiScreenItemData_8" at 469,45 size 355x40; TextOn 'Back'; TextOff 'Text'
   TextField "Screen title" at 455,41 size 373x50; Text 'Screen title'

screen "RIO 01 Digital Inputs" 1280x800, template "Template"
   on GenerateScreen: "TitleUpdater"()
   TextField "Text field_37" at 16,52 size 476x26; Text 'RIO #1 (Remote Inputs & Outputs Panel No. 1)'
   TextField "Text field_38" at 16,122 size 55x22; Text 'I0.0'
   TextField "Text field_39" at 16,157 size 55x22; Text 'I0.1'
   TextField "Text field_40" at 16,193 size 55x22; Text 'I0.2'
   TextField "Text field_41" at 16,229 size 55x22; Text 'I0.3'
   TextField "Text field_42" at 16,265 size 55x22; Text 'I0.4'
   TextField "Text field_43" at 16,301 size 55x22; Text 'I0.5'
   TextField "Text field_44" at 16,337 size 55x22; Text 'I0.6'
   TextField "Text field_45" at 16,373 size 55x22; Text 'I0.7'
   Circle "Circle_33" at 76,123 size 20x20
      Appearance <- "FPT GTT Isolation Valve Feedback - Opened"
   Circle "Circle_34" at 76,158 size 20x20
      Appearance <- "FPT GTT Isolation Valve Feedback - Closed"
   Circle "Circle_35" at 76,194 size 20x20
      Appearance <- "FPT Tank Vent Valve 1 Feedback - Opened"
   Circle "Circle_36" at 76,230 size 20x20
      Appearance <- "FPT Tank Vent Valve 1 Feedback - Closed"
   Circle "Circle_37" at 76,265 size 20x20
      Appearance <- "FPT Tank Vent Valve 2 Feedback - Opened"
   Circle "Circle_38" at 76,301 size 20x20
      Appearance <- "FPT Tank Vent Valve 2 Feedback - Closed"
   Circle "Circle_39" at 76,337 size 20x20
      Appearance <- "RIO1_SPR_DI_0_6"
   Circle "Circle_40" at 76,373 size 20x20
      Appearance <- "RIO1_SPR_DI_0_7"
   TextField "Text field_46" at 33,90 size 49x26; Text 'I0'
   TextField "Text field_47" at 16,441 size 55x22; Text 'I3.0'
   TextField "Text field_48" at 16,476 size 55x22; Text 'I3.1'
   TextField "Text field_49" at 16,512 size 55x22; Text 'I3.2'
   TextField "Text field_50" at 16,548 size 55x22; Text 'I3.3'
   TextField "Text field_51" at 16,584 size 55x22; Text 'I3.4'
   TextField "Text field_52" at 16,620 size 55x22; Text 'I3.5'
   TextField "Text field_53" at 16,656 size 55x22; Text 'I3.6'
   TextField "Text field_54" at 16,692 size 55x22; Text 'I3.7'
   Circle "Circle_41" at 76,442 size 20x20
      Appearance <- "Tank 1P GTT Isolation Valve Feedback - Opened"
   Circle "Circle_42" at 76,477 size 20x20
      Appearance <- "Tank 1P GTT Isolation Valve Feedback - Closed"
   Circle "Circle_43" at 76,513 size 20x20
      Appearance <- "Tank 1P Tank Vent Valve 1 Feedback - Opened"
   Circle "Circle_44" at 76,549 size 20x20
      Appearance <- "Tank 1P Tank Vent Valve 1 Feedback - Closed"
   Circle "Circle_45" at 76,585 size 20x20
      Appearance <- "Tank 1P Tank Vent Valve 2 Feedback - Opened"
   Circle "Circle_46" at 76,621 size 20x20
      Appearance <- "Tank 1P Tank Vent Valve 2 Feedback - Closed"
   Circle "Circle_47" at 76,657 size 20x20
      Appearance <- "RIO1_SPR_DI_3_6"
   Circle "Circle_48" at 76,693 size 20x20
      Appearance <- "RIO1_SPR_DI_3_7"
   TextField "Text field_55" at 33,409 size 49x26; Text 'I1'
   TextField "Text field_56" at 548,122 size 55x22; Text 'I6.0'
   TextField "Text field_57" at 548,157 size 55x22; Text 'I6.1'
   TextField "Text field_58" at 548,193 size 55x22; Text 'I6.2'
   TextField "Text field_59" at 548,229 size 55x22; Text 'I6.3'
   TextField "Text field_60" at 548,265 size 55x22; Text 'I6.4'
   TextField "Text field_61" at 548,301 size 55x22; Text 'I6.5'
   TextField "Text field_62" at 548,337 size 55x22; Text 'I6.6'
   TextField "Text field_63" at 548,373 size 55x22; Text 'I6.7'
   Circle "Circle_49" at 608,122 size 20x20
      Appearance <- "Tank 1S GTT Isolation Valve Feedback - Opened"
   Circle "Circle_50" at 608,157 size 20x20
      Appearance <- "Tank 1S GTT Isolation Valve Feedback - Closed"
   Circle "Circle_51" at 608,193 size 20x20
      Appearance <- "Tank 1S Tank Vent Valve 1 Feedback - Opened"
   Circle "Circle_52" at 608,229 size 20x20
      Appearance <- "Tank 1S Tank Vent Valve 1 Feedback - Closed"
   Circle "Circle_53" at 608,265 size 20x20
      Appearance <- "Tank 1S Tank Vent Valve 2 Feedback - Opened"
   Circle "Circle_54" at 608,301 size 20x20
      Appearance <- "Tank 1S Tank Vent Valve 2 Feedback - Closed"
   Circle "Circle_55" at 608,337 size 20x20
      Appearance <- "RIO1_SPR_DI_6_6"
   Circle "Circle_56" at 608,373 size 20x20
      Appearance <- "RIO1_SPR_DI_6_7"
   TextField "Text field_64" at 570,90 size 49x26; Text 'I2'
   TextField "Text field_65" at 546,441 size 46x22; Text 'I9.0'
   TextField "Text field_66" at 546,476 size 46x22; Text 'I9.1'
   TextField "Text field_67" at 546,512 size 46x22; Text 'I9.2'
   TextField "Text field_68" at 546,548 size 46x22; Text 'I9.3'
   TextField "Text field_69" at 546,584 size 46x22; Text 'I9.4'
   TextField "Text field_70" at 546,620 size 46x22; Text 'I9.5'
   TextField "Text field_71" at 546,656 size 46x22; Text 'I9.6'
   TextField "Text field_72" at 546,692 size 46x22; Text 'I9.7'
   Circle "Circle_57" at 606,441 size 20x20
      Appearance <- "FPT BWT Level High High Switch"
   Circle "Circle_58" at 606,476 size 20x20
      Appearance <- "RIO1 Tanks Pressure Switch Hi Hi"
   Circle "Circle_59" at 606,512 size 20x20
      Appearance <- "Tank 1P BWT Level High High Switch"
   Circle "Circle_60" at 606,548 size 20x20
      Appearance <- "Tank 1S BWT Level High High Switch"
   Circle "Circle_61" at 606,584 size 20x20
      Appearance <- "RIO1_SPR_DI_9_4"
   Circle "Circle_62" at 606,620 size 20x20
      Appearance <- "RIO1_SPR_DI_9_5"
   Circle "Circle_63" at 606,656 size 20x20
      Appearance <- "RIO1_SPR_DI_9_6"
   Circle "Circle_64" at 606,692 size 20x20
      Appearance <- "RIO1_SPR_DI_9_7"
   TextField "Text field_73" at 563,409 size 49x26; Text 'I3'
   Button "HmiScreenItemData_1" at 1,1 size 150x43; TextOn 'Back'; TextOff 'Commissioning'
      on Release: ActivateScreen("Commissioning Main Page", 0)
   TextField "Text field_107" at 105,114 size 348x38; Text 'FPT GTT Isolation Valve Feedback - Opened CV422'
   TextField "Text field_108" at 105,149 size 340x38; Text 'FPT GTT Isolation Valve Feedback - Closed CV422'
   TextField "Text field_109" at 105,184 size 337x38; Text 'FPT Tank Vent Valve 1 Feedback - Opened CV441-FPTA'
   TextField "Text field_110" at 105,220 size 329x38; Text 'FPT Tank Vent Valve 1 Feedback - Closed CV441-FPTA'
   TextField "Text field_111" at 105,255 size 337x38; Text 'FPT Tank Vent Valve 2 Feedback - Opened CV441-FPTB'
   TextField "Text field_112" at 105,291 size 329x38; Text 'FPT Tank Vent Valve 2 Feedback - Closed CV441-FPTB'
   TextField "Text field_113" at 104,328 size 100x21; Text 'Spare Input'
   TextField "Text field_114" at 104,365 size 100x21; Text 'Spare Input'